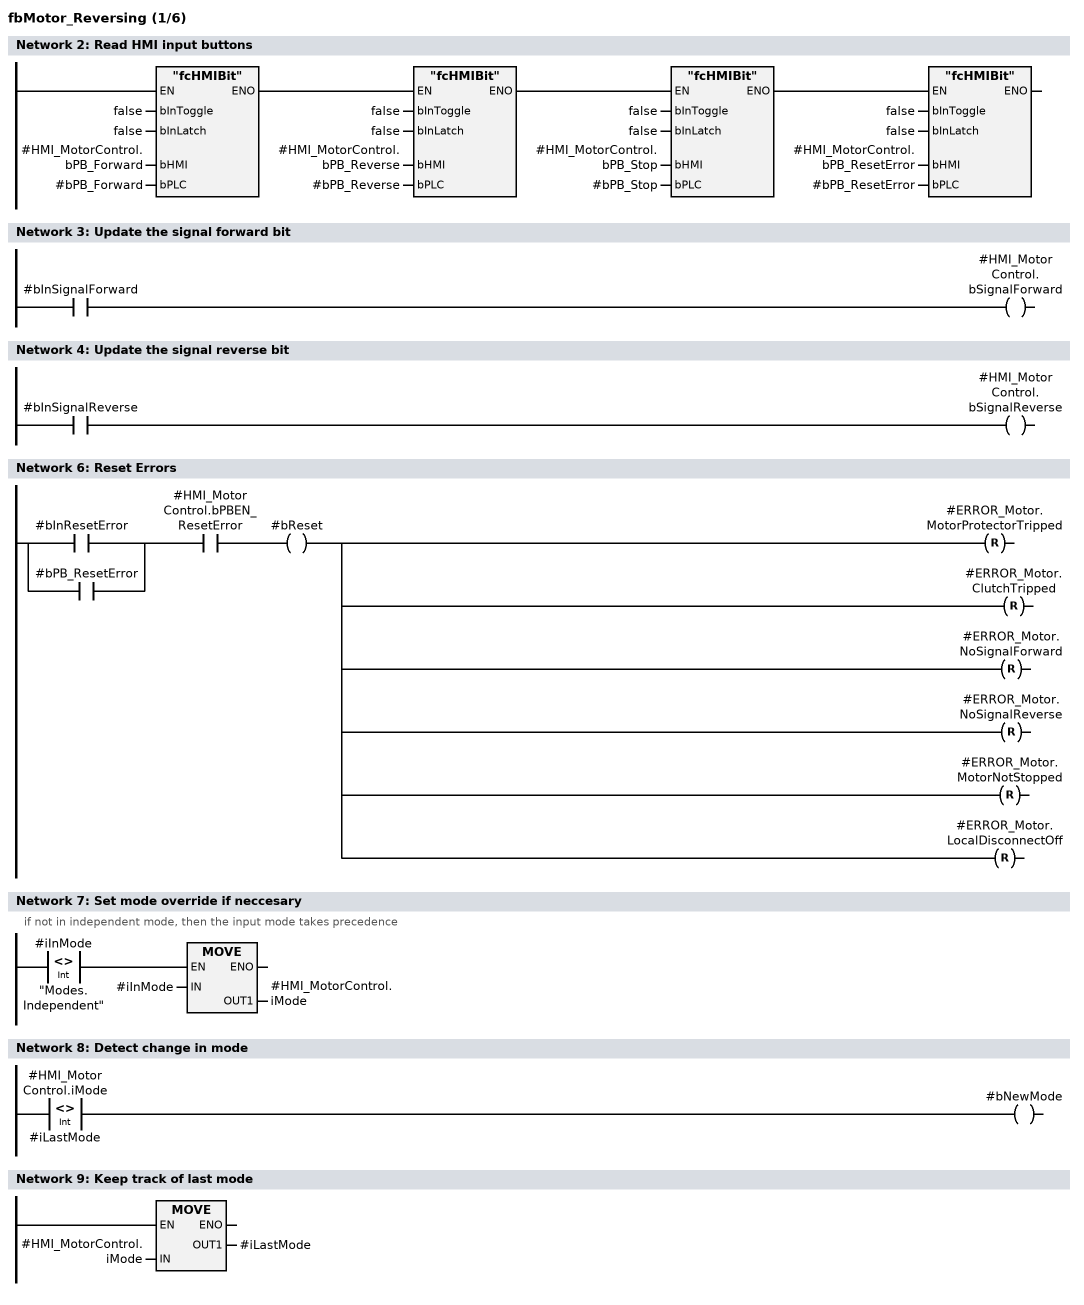
   RUNG wire#powerrail
      "fcHMIBit"(bInToggle := false, bInLatch := false, bHMI := #HMI_MotorControl.bPB_Forward, bPLC := #bPB_Forward)
      "fcHMIBit"(bInToggle := false, bInLatch := false, bHMI := #HMI_MotorControl.bPB_Reverse, bPLC := #bPB_Reverse)
      "fcHMIBit"(bInToggle := false, bInLatch := false, bHMI := #HMI_MotorControl.bPB_Stop, bPLC := #bPB_Stop)
      "fcHMIBit"(bInToggle := false, bInLatch := false, bHMI := #HMI_MotorControl.bPB_ResetError, bPLC := #bPB_ResetError)
   END_RUNG
   // the same network as SCL:
   "fcHMIBit"(bInToggle := false,
              bInLatch := false,
              bHMI := #HMI_MotorControl.bPB_Forward,
              bPLC := #bPB_Forward,
              ENO => #_w1);
   "fcHMIBit"(EN := #_w1,
              bInToggle := false,
              bInLatch := false,
              bHMI := #HMI_MotorControl.bPB_Reverse,
              bPLC := #bPB_Reverse,
              ENO => #_w2);
   "fcHMIBit"(EN := #_w2,
              bInToggle := false,
              bInLatch := false,
              bHMI := #HMI_MotorControl.bPB_Stop,
              bPLC := #bPB_Stop,
              ENO => #_w3);
   IF #_w3 THEN
       "fcHMIBit"(bInToggle := false,
                  bInLatch := false,
                  bHMI := #HMI_MotorControl.bPB_ResetError,
                  bPLC := #bPB_ResetError);
   END_IF;
END_REGION

REGION Network 3: Update the signal forward bit
   RUNG wire#powerrail
      Contact( #bInSignalForward )
      Coil( #HMI_MotorControl.bSignalForward )
   END_RUNG
   // the same network as SCL:
   #HMI_MotorControl.bSignalForward := #bInSignalForward;
END_REGION

REGION Network 4: Update the signal reverse bit
   RUNG wire#powerrail
      Contact( #bInSignalReverse )
      Coil( #HMI_MotorControl.bSignalReverse )
   END_RUNG
   // the same network as SCL:
   #HMI_MotorControl.bSignalReverse := #bInSignalReverse;
END_REGION

REGION Network 5: --------------------------------------------------- Control Logic ------------------------------------------------------------
END_REGION

REGION Network 6: Reset Errors
   RUNG wire#powerrail
      Contact( #bInResetError )
      wire#w1
      Contact( #HMI_MotorControl.bPBEN_ResetError )
      Coil( #bReset )
      wire#w2
      R_Coil( #ERROR_Motor.MotorProtectorTripped )
   END_RUNG
   RUNG wire#powerrail
      Contact( #bPB_ResetError )
   END_RUNG wire#w1
   RUNG wire#w2
      R_Coil( #ERROR_Motor.ClutchTripped )
   END_RUNG
   RUNG wire#w2
      R_Coil( #ERROR_Motor.NoSignalForward )
   END_RUNG
   RUNG wire#w2
      R_Coil( #ERROR_Motor.NoSignalReverse )
   END_RUNG
   RUNG wire#w2
      R_Coil( #ERROR_Motor.MotorNotStopped )
   END_RUNG
   RUNG wire#w2
      R_Coil( #ERROR_Motor.LocalDisconnectOff )
   END_RUNG
   // the same network as SCL:
   #bReset := (#bInResetError OR #bPB_ResetError) AND #HMI_MotorControl.bPBEN_ResetError;
   IF #bReset THEN
       #ERROR_Motor.MotorProtectorTripped := FALSE;
       #ERROR_Motor.ClutchTripped := FALSE;
       #ERROR_Motor.NoSignalForward := FALSE;
       #ERROR_Motor.NoSignalReverse := FALSE;
       #ERROR_Motor.MotorNotStopped := FALSE;
       #ERROR_Motor.LocalDisconnectOff := FALSE;
   END_IF;
END_REGION

REGION Network 7: Set mode override if neccesary
   // if not in independent mode, then the input mode takes precedence
   RUNG wire#powerrail
      { S7_Templates := "SrcType := Int" } NE_Contact(in1 := #iInMode, in2 := "Modes.Independent")
      { S7_GenerateENO := "TRUE" } Move(in := #iInMode, out1 => #HMI_MotorControl.iMode)
   END_RUNG
   // the same network as SCL:
   IF #iInMode <> "Modes.Independent" THEN #HMI_MotorControl.iMode := #iInMode; END_IF;
END_REGION

REGION Network 8: Detect change in mode
   RUNG wire#powerrail
      { S7_Templates := "SrcType := Int" } NE_Contact(in1 := #HMI_MotorControl.iMode, in2 := #iLastMode)
      Coil( #bNewMode )
   END_RUNG
   // the same network as SCL:
   #bNewMode := #HMI_MotorControl.iMode <> #iLastMode;
END_REGION

REGION Network 9: Keep track of last mode
   RUNG wire#powerrail
      { S7_GenerateENO := "TRUE" } Move(in := #HMI_MotorControl.iMode, out1 => #iLastMode)
   END_RUNG
   // the same network as SCL:
   #iLastMode := #HMI_MotorControl.iMode;
END_REGION

REGION Network 10: Determine if auto or manual mode is active
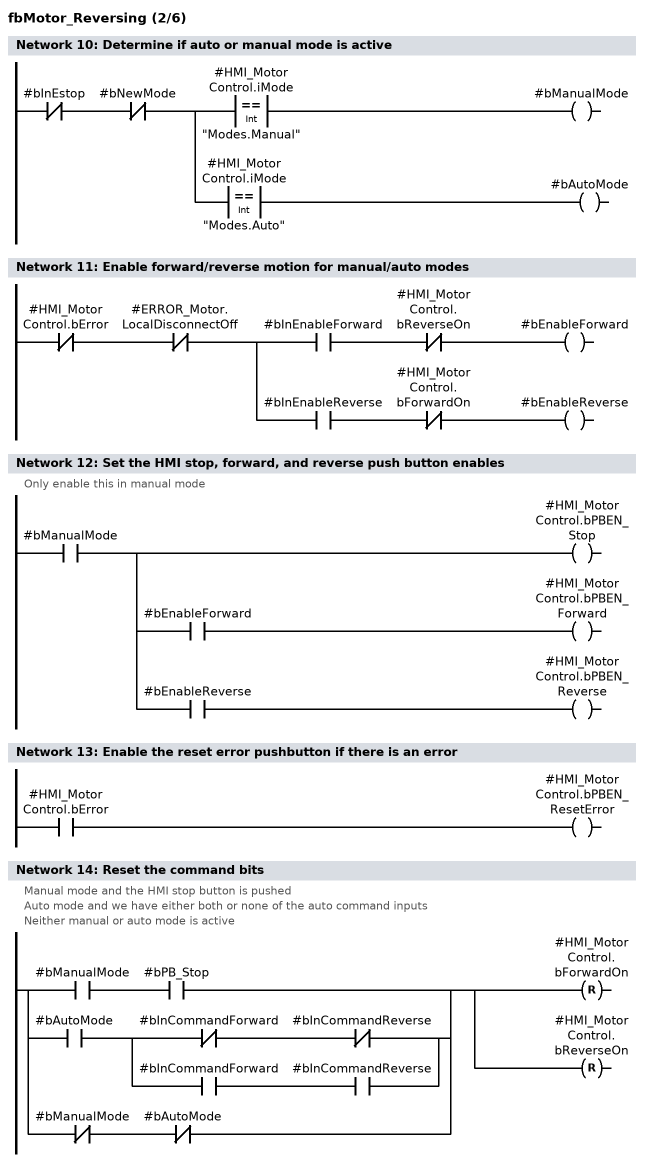
   RUNG wire#powerrail
      I_Contact( #bInEstop )
      I_Contact( #bNewMode )
      wire#w1
      { S7_Templates := "SrcType := Int" } EQ_Contact(in1 := #HMI_MotorControl.iMode, in2 := "Modes.Manual")
      Coil( #bManualMode )
   END_RUNG
   RUNG wire#w1
      { S7_Templates := "SrcType := Int" } EQ_Contact(in1 := #HMI_MotorControl.iMode, in2 := "Modes.Auto")
      Coil( #bAutoMode )
   END_RUNG
   // the same network as SCL:
   #_w1 := NOT #bInEstop AND NOT #bNewMode;
   #bManualMode := #_w1 AND (#HMI_MotorControl.iMode = "Modes.Manual");
   #bAutoMode := #_w1 AND (#HMI_MotorControl.iMode = "Modes.Auto");
END_REGION

REGION Network 11: Enable forward/reverse motion for manual/auto modes
   RUNG wire#powerrail
      I_Contact( #HMI_MotorControl.bError )
      I_Contact( #ERROR_Motor.LocalDisconnectOff )
      wire#w1
      Contact( #bInEnableForward )
      I_Contact( #HMI_MotorControl.bReverseOn )
      Coil( #bEnableForward )
   END_RUNG
   RUNG wire#w1
      Contact( #bInEnableReverse )
      I_Contact( #HMI_MotorControl.bForwardOn )
      Coil( #bEnableReverse )
   END_RUNG
   // the same network as SCL:
   #_w1 := NOT #HMI_MotorControl.bError AND NOT #ERROR_Motor.LocalDisconnectOff;
   #bEnableForward := #_w1 AND #bInEnableForward AND NOT #HMI_MotorControl.bReverseOn;
   #bEnableReverse := #_w1 AND #bInEnableReverse AND NOT #HMI_MotorControl.bForwardOn;
END_REGION

REGION Network 12: Set the HMI stop, forward, and reverse push button enables
   // Only enable this in manual mode
   RUNG wire#powerrail
      Contact( #bManualMode )
      wire#w1
      Coil( #HMI_MotorControl.bPBEN_Stop )
   END_RUNG
   RUNG wire#w1
      Contact( #bEnableForward )
      Coil( #HMI_MotorControl.bPBEN_Forward )
   END_RUNG
   RUNG wire#w1
      Contact( #bEnableReverse )
      Coil( #HMI_MotorControl.bPBEN_Reverse )
   END_RUNG
   // the same network as SCL:
   #HMI_MotorControl.bPBEN_Stop := #bManualMode;
   #HMI_MotorControl.bPBEN_Forward := #bManualMode AND #bEnableForward;
   #HMI_MotorControl.bPBEN_Reverse := #bManualMode AND #bEnableReverse;
END_REGION

REGION Network 13: Enable the reset error pushbutton if there is an error
   RUNG wire#powerrail
      Contact( #HMI_MotorControl.bError )
      Coil( #HMI_MotorControl.bPBEN_ResetError )
   END_RUNG
   // the same network as SCL:
   #HMI_MotorControl.bPBEN_ResetError := #HMI_MotorControl.bError;
END_REGION

REGION Network 14: Reset the command bits
   // Manual mode and the HMI stop button is pushed
   // Auto mode and we have either both or none of the auto command inputs
   // Neither manual or auto mode is active
   RUNG wire#powerrail
      Contact( #bManualMode )
      Contact( #bPB_Stop )
      wire#w1
      R_Coil( #HMI_MotorControl.bForwardOn )
   END_RUNG
   RUNG wire#powerrail
      Contact( #bAutoMode )
      wire#w2
      I_Contact( #bInCommandForward )
      I_Contact( #bInCommandReverse )
   END_RUNG wire#w1
   RUNG wire#w2
      Contact( #bInCommandForward )
      Contact( #bInCommandReverse )
   END_RUNG wire#w1
   RUNG wire#powerrail
      I_Contact( #bManualMode )
      I_Contact( #bAutoMode )
   END_RUNG wire#w1
   RUNG wire#w1
      R_Coil( #HMI_MotorControl.bReverseOn )
   END_RUNG
   // the same network as SCL:
   IF (#bManualMode AND #bPB_Stop) OR (#bAutoMode AND ((NOT #bInCommandForward AND NOT #bInCommandReverse) OR (#bInCommandForward AND #bInCommandReverse))) OR (NOT #bManualMode AND NOT #bAutoMode) THEN
       #HMI_MotorControl.bForwardOn := FALSE;
       #HMI_MotorControl.bReverseOn := FALSE;
   END_IF;
END_REGION

REGION Network 15: Start forward request
   // Manual mode and only a start forward button is pressed and enabled
   // Auto mode when we receive a auto command and it is enabled
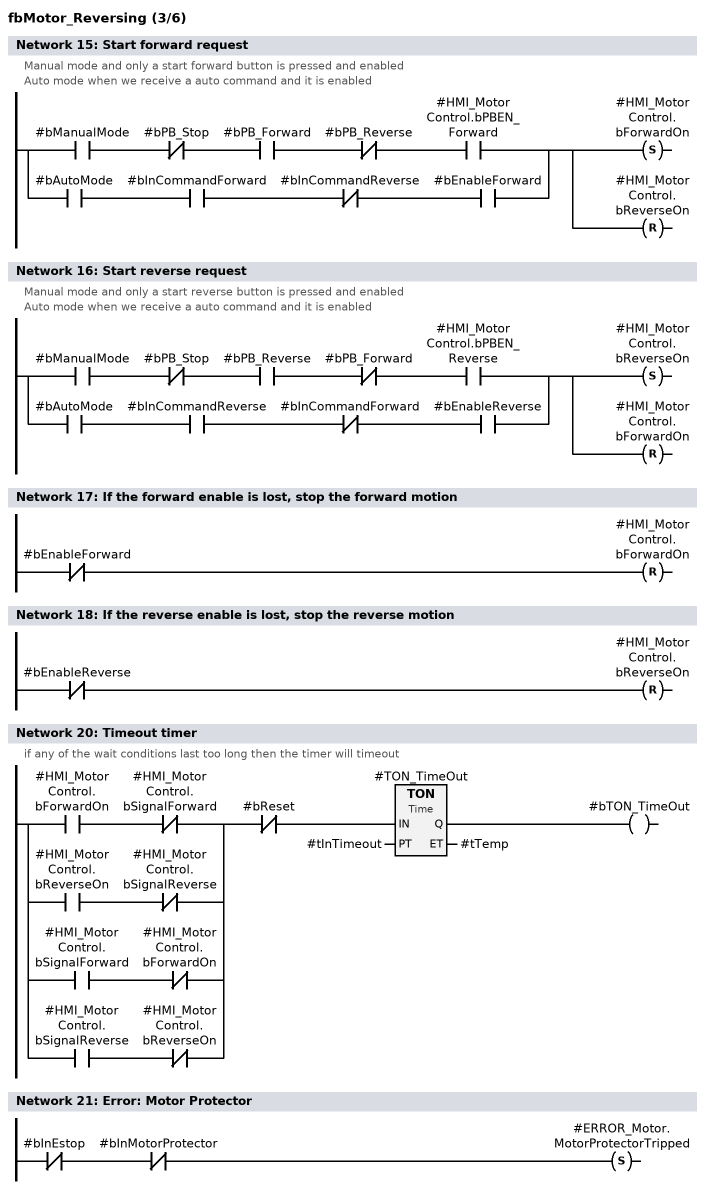
   RUNG wire#powerrail
      Contact( #bManualMode )
      I_Contact( #bPB_Stop )
      Contact( #bPB_Forward )
      I_Contact( #bPB_Reverse )
      Contact( #HMI_MotorControl.bPBEN_Forward )
      wire#w1
      S_Coil( #HMI_MotorControl.bForwardOn )
   END_RUNG
   RUNG wire#powerrail
      Contact( #bAutoMode )
      Contact( #bInCommandForward )
      I_Contact( #bInCommandReverse )
      Contact( #bEnableForward )
   END_RUNG wire#w1
   RUNG wire#w1
      R_Coil( #HMI_MotorControl.bReverseOn )
   END_RUNG
   // the same network as SCL:
   IF (#bManualMode AND NOT #bPB_Stop AND #bPB_Forward AND NOT #bPB_Reverse AND #HMI_MotorControl.bPBEN_Forward) OR (#bAutoMode AND #bInCommandForward AND NOT #bInCommandReverse AND #bEnableForward) THEN
       #HMI_MotorControl.bForwardOn := TRUE;
       #HMI_MotorControl.bReverseOn := FALSE;
   END_IF;
END_REGION

REGION Network 16: Start reverse request
   // Manual mode and only a start reverse button is pressed and enabled
   // Auto mode when we receive a auto command and it is enabled
   RUNG wire#powerrail
      Contact( #bManualMode )
      I_Contact( #bPB_Stop )
      Contact( #bPB_Reverse )
      I_Contact( #bPB_Forward )
      Contact( #HMI_MotorControl.bPBEN_Reverse )
      wire#w1
      S_Coil( #HMI_MotorControl.bReverseOn )
   END_RUNG
   RUNG wire#powerrail
      Contact( #bAutoMode )
      Contact( #bInCommandReverse )
      I_Contact( #bInCommandForward )
      Contact( #bEnableReverse )
   END_RUNG wire#w1
   RUNG wire#w1
      R_Coil( #HMI_MotorControl.bForwardOn )
   END_RUNG
   // the same network as SCL:
   IF (#bManualMode AND NOT #bPB_Stop AND #bPB_Reverse AND NOT #bPB_Forward AND #HMI_MotorControl.bPBEN_Reverse) OR (#bAutoMode AND #bInCommandReverse AND NOT #bInCommandForward AND #bEnableReverse) THEN
       #HMI_MotorControl.bReverseOn := TRUE;
       #HMI_MotorControl.bForwardOn := FALSE;
   END_IF;
END_REGION

REGION Network 17: If the forward enable is lost, stop the forward motion
   RUNG wire#powerrail
      I_Contact( #bEnableForward )
      R_Coil( #HMI_MotorControl.bForwardOn )
   END_RUNG
   // the same network as SCL:
   IF NOT #bEnableForward THEN #HMI_MotorControl.bForwardOn := FALSE; END_IF;
END_REGION

REGION Network 18: If the reverse enable is lost, stop the reverse motion
   RUNG wire#powerrail
      I_Contact( #bEnableReverse )
      R_Coil( #HMI_MotorControl.bReverseOn )
   END_RUNG
   // the same network as SCL:
   IF NOT #bEnableReverse THEN #HMI_MotorControl.bReverseOn := FALSE; END_IF;
END_REGION

REGION Network 19: --------------------------------------------------------- Errors ------------------------------------------------------------------
END_REGION

REGION Network 20: Timeout timer
   // if any of the wait conditions last too long then the timer will timeout
   #TON_TimeOut.TON(IN := ((#HMI_MotorControl.bForwardOn AND NOT #HMI_MotorControl.bSignalForward) OR (#HMI_MotorControl.bReverseOn AND NOT #HMI_MotorControl.bSignalReverse) OR (#HMI_MotorControl.bSignalForward AND NOT #HMI_MotorControl.bForwardOn) OR (#HMI_MotorControl.bSignalReverse AND NOT #HMI_MotorControl.bReverseOn)) AND NOT #bReset,
                    PT := #tInTimeout,
                    ET => #tTemp);
   #bTON_TimeOut := #TON_TimeOut.Q;
END_REGION

REGION Network 21: Error: Motor Protector
   RUNG wire#powerrail
      I_Contact( #bInEstop )
      I_Contact( #bInMotorProtector )
      S_Coil( #ERROR_Motor.MotorProtectorTripped )
   END_RUNG
   // the same network as SCL:
   IF NOT #bInEstop AND NOT #bInMotorProtector THEN #ERROR_Motor.MotorProtectorTripped := TRUE; END_IF;
END_REGION

REGION Network 22: Error: Kill Switch/ local disconnect
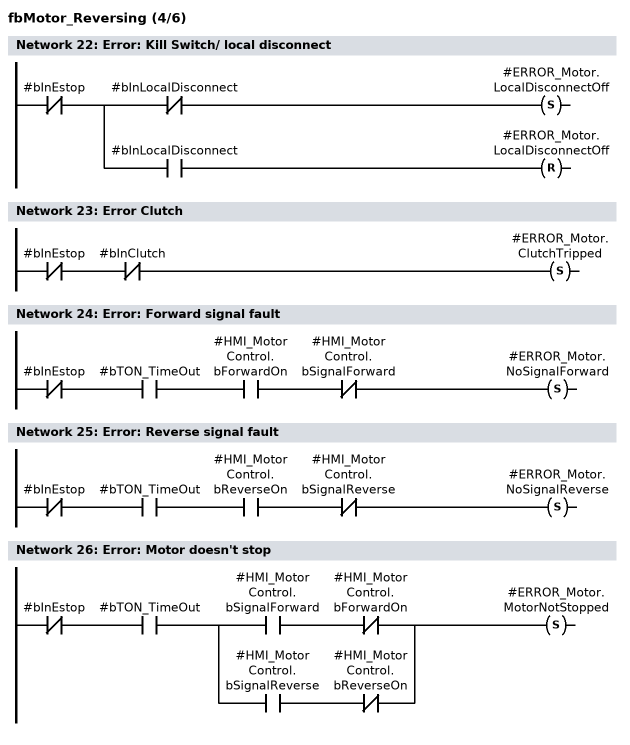
   RUNG wire#powerrail
      I_Contact( #bInEstop )
      wire#w1
      I_Contact( #bInLocalDisconnect )
      S_Coil( #ERROR_Motor.LocalDisconnectOff )
   END_RUNG
   RUNG wire#w1
      Contact( #bInLocalDisconnect )
      R_Coil( #ERROR_Motor.LocalDisconnectOff )
   END_RUNG
   // the same network as SCL:
   IF NOT #bInEstop AND NOT #bInLocalDisconnect THEN #ERROR_Motor.LocalDisconnectOff := TRUE; END_IF;
   IF NOT #bInEstop AND #bInLocalDisconnect THEN #ERROR_Motor.LocalDisconnectOff := FALSE; END_IF;
END_REGION

REGION Network 23: Error Clutch
   RUNG wire#powerrail
      I_Contact( #bInEstop )
      I_Contact( #bInClutch )
      S_Coil( #ERROR_Motor.ClutchTripped )
   END_RUNG
   // the same network as SCL:
   IF NOT #bInEstop AND NOT #bInClutch THEN #ERROR_Motor.ClutchTripped := TRUE; END_IF;
END_REGION

REGION Network 24: Error: Forward signal fault
   RUNG wire#powerrail
      I_Contact( #bInEstop )
      Contact( #bTON_TimeOut )
      Contact( #HMI_MotorControl.bForwardOn )
      I_Contact( #HMI_MotorControl.bSignalForward )
      S_Coil( #ERROR_Motor.NoSignalForward )
   END_RUNG
   // the same network as SCL:
   IF NOT #bInEstop AND #bTON_TimeOut AND #HMI_MotorControl.bForwardOn AND NOT #HMI_MotorControl.bSignalForward THEN
       #ERROR_Motor.NoSignalForward := TRUE;
   END_IF;
END_REGION

REGION Network 25: Error: Reverse signal fault
   RUNG wire#powerrail
      I_Contact( #bInEstop )
      Contact( #bTON_TimeOut )
      Contact( #HMI_MotorControl.bReverseOn )
      I_Contact( #HMI_MotorControl.bSignalReverse )
      S_Coil( #ERROR_Motor.NoSignalReverse )
   END_RUNG
   // the same network as SCL:
   IF NOT #bInEstop AND #bTON_TimeOut AND #HMI_MotorControl.bReverseOn AND NOT #HMI_MotorControl.bSignalReverse THEN
       #ERROR_Motor.NoSignalReverse := TRUE;
   END_IF;
END_REGION

REGION Network 26: Error: Motor doesn't stop
   RUNG wire#powerrail
      I_Contact( #bInEstop )
      Contact( #bTON_TimeOut )
      wire#w1
      Contact( #HMI_MotorControl.bSignalForward )
      I_Contact( #HMI_MotorControl.bForwardOn )
      wire#w2
      S_Coil( #ERROR_Motor.MotorNotStopped )
   END_RUNG
   RUNG wire#w1
      Contact( #HMI_MotorControl.bSignalReverse )
      I_Contact( #HMI_MotorControl.bReverseOn )
   END_RUNG wire#w2
   // the same network as SCL:
   IF NOT #bInEstop AND #bTON_TimeOut AND ((#HMI_MotorControl.bSignalForward AND NOT #HMI_MotorControl.bForwardOn) OR (#HMI_MotorControl.bSignalReverse AND NOT #HMI_MotorControl.bReverseOn)) THEN
       #ERROR_Motor.MotorNotStopped := TRUE;
   END_IF;
END_REGION

REGION Network 27: Scroll errors on the HMI
   // This block loops through all of the possible erros and displays them on the HMI 
   // by setting an index value for each error bit.
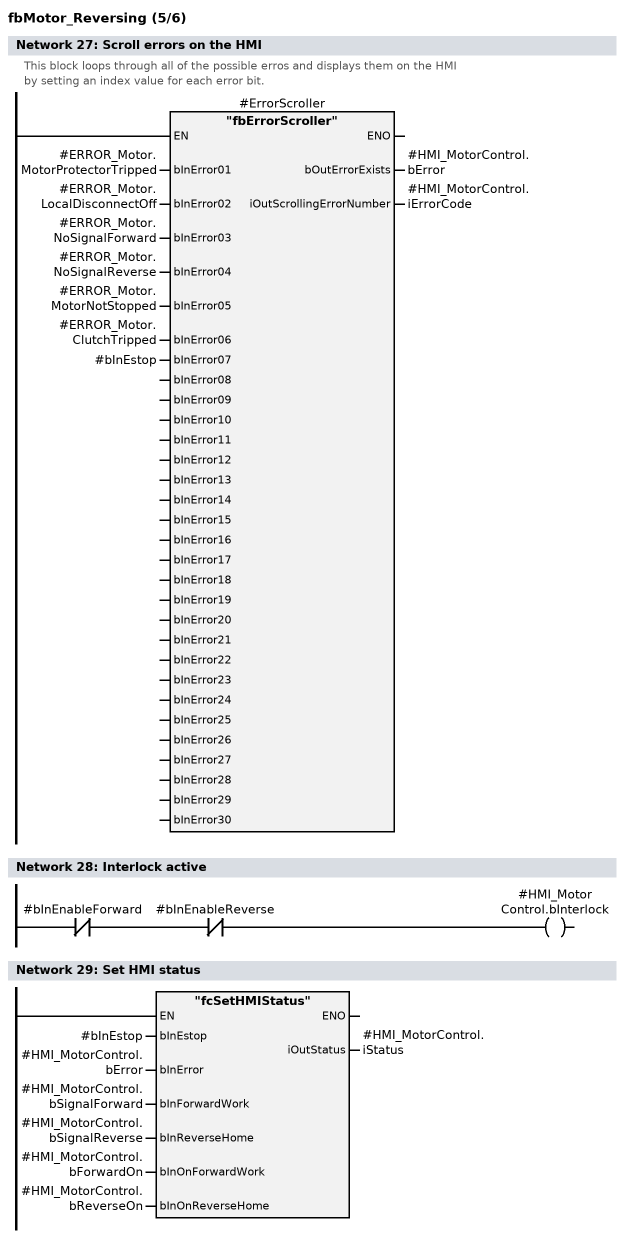
   RUNG wire#powerrail
      #ErrorScroller(bInError01 := #ERROR_Motor.MotorProtectorTripped, bInError02 := #ERROR_Motor.LocalDisconnectOff, bInError03 := #ERROR_Motor.NoSignalForward, bInError04 := #ERROR_Motor.NoSignalReverse, bInError05 := #ERROR_Motor.MotorNotStopped, bInError06 := #ERROR_Motor.ClutchTripped, bInError07 := #bInEstop, bInError08 :=, bInError09 :=, bInError10 :=, bInError11 :=, bInError12 :=, bInError13 :=, bInError14 :=, bInError15 :=, bInError16 :=, bInError17 :=, bInError18 :=, bInError19 :=, bInError20 :=, bInError21 :=, bInError22 :=, bInError23 :=, bInError24 :=, bInError25 :=, bInError26 :=, bInError27 :=, bInError28 :=, bInError29 :=, bInError30 :=, bOutErrorExists => #HMI_MotorControl.bError, iOutScrollingErrorNumber => #HMI_MotorControl.iErrorCode)
   END_RUNG
   // the same network as SCL:
   #ErrorScroller(bInError01 := #ERROR_Motor.MotorProtectorTripped,   // "fbErrorScroller"
                  bInError02 := #ERROR_Motor.LocalDisconnectOff,
                  bInError03 := #ERROR_Motor.NoSignalForward,
                  bInError04 := #ERROR_Motor.NoSignalReverse,
                  bInError05 := #ERROR_Motor.MotorNotStopped,
                  bInError06 := #ERROR_Motor.ClutchTripped,
                  bInError07 := #bInEstop,
                  bOutErrorExists => #HMI_MotorControl.bError,
                  iOutScrollingErrorNumber => #HMI_MotorControl.iErrorCode);
END_REGION

REGION Network 28: Interlock active
   RUNG wire#powerrail
      I_Contact( #bInEnableForward )
      I_Contact( #bInEnableReverse )
      Coil( #HMI_MotorControl.bInterlock )
   END_RUNG
   // the same network as SCL:
   #HMI_MotorControl.bInterlock := NOT #bInEnableForward AND NOT #bInEnableReverse;
END_REGION

REGION Network 29: Set HMI status
   RUNG wire#powerrail
      "fcSetHMIStatus"(bInEstop := #bInEstop, bInError := #HMI_MotorControl.bError, bInForwardWork := #HMI_MotorControl.bSignalForward, bInReverseHome := #HMI_MotorControl.bSignalReverse, bInOnForwardWork := #HMI_MotorControl.bForwardOn, bInOnReverseHome := #HMI_MotorControl.bReverseOn, iOutStatus => #HMI_MotorControl.iStatus)
   END_RUNG
   // the same network as SCL:
   "fcSetHMIStatus"(bInEstop := #bInEstop,
                    bInError := #HMI_MotorControl.bError,
                    bInForwardWork := #HMI_MotorControl.bSignalForward,
                    bInReverseHome := #HMI_MotorControl.bSignalReverse,
                    bInOnForwardWork := #HMI_MotorControl.bForwardOn,
                    bInOnReverseHome := #HMI_MotorControl.bReverseOn,
                    iOutStatus => #HMI_MotorControl.iStatus);
END_REGION

REGION Network 30: ------------------------------------------------- Outputs --------------------------------------------------
END_REGION

REGION Network 31: Output: Forward
   // Forward
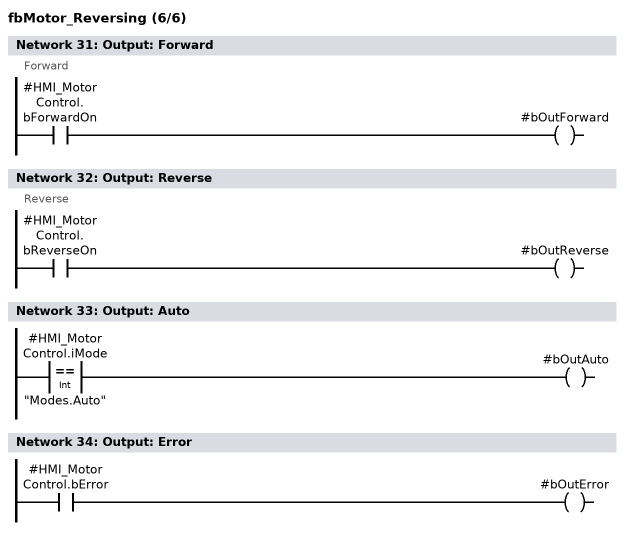
   RUNG wire#powerrail
      Contact( #HMI_MotorControl.bForwardOn )
      Coil( #bOutForward )
   END_RUNG
   // the same network as SCL:
   #bOutForward := #HMI_MotorControl.bForwardOn;
END_REGION

REGION Network 32: Output: Reverse
   // Reverse
   RUNG wire#powerrail
      Contact( #HMI_MotorControl.bReverseOn )
      Coil( #bOutReverse )
   END_RUNG
   // the same network as SCL:
   #bOutReverse := #HMI_MotorControl.bReverseOn;
END_REGION

REGION Network 33: Output: Auto
   RUNG wire#powerrail
      { S7_Templates := "SrcType := Int" } EQ_Contact(in1 := #HMI_MotorControl.iMode, in2 := "Modes.Auto")
      Coil( #bOutAuto )
   END_RUNG
   // the same network as SCL:
   #bOutAuto := #HMI_MotorControl.iMode = "Modes.Auto";
END_REGION

REGION Network 34: Output: Error
   RUNG wire#powerrail
      Contact( #HMI_MotorControl.bError )
      Coil( #bOutError )
   END_RUNG
   // the same network as SCL:
   #bOutError := #HMI_MotorControl.bError;
END_REGION
END_FUNCTION_BLOCK

FUNCTION_BLOCK "fbIO_AnalogInput"   // FB140, LAD
TITLE = Reads and controls an analog input
{ S7_Optimized_Access := 'FALSE' }
VERSION : 0.1
BEGIN

REGION Network 1: --------------------------------------------------------- Inputs ------------------------------------------------------------------
END_REGION

REGION Network 2: Read HMI input buttons
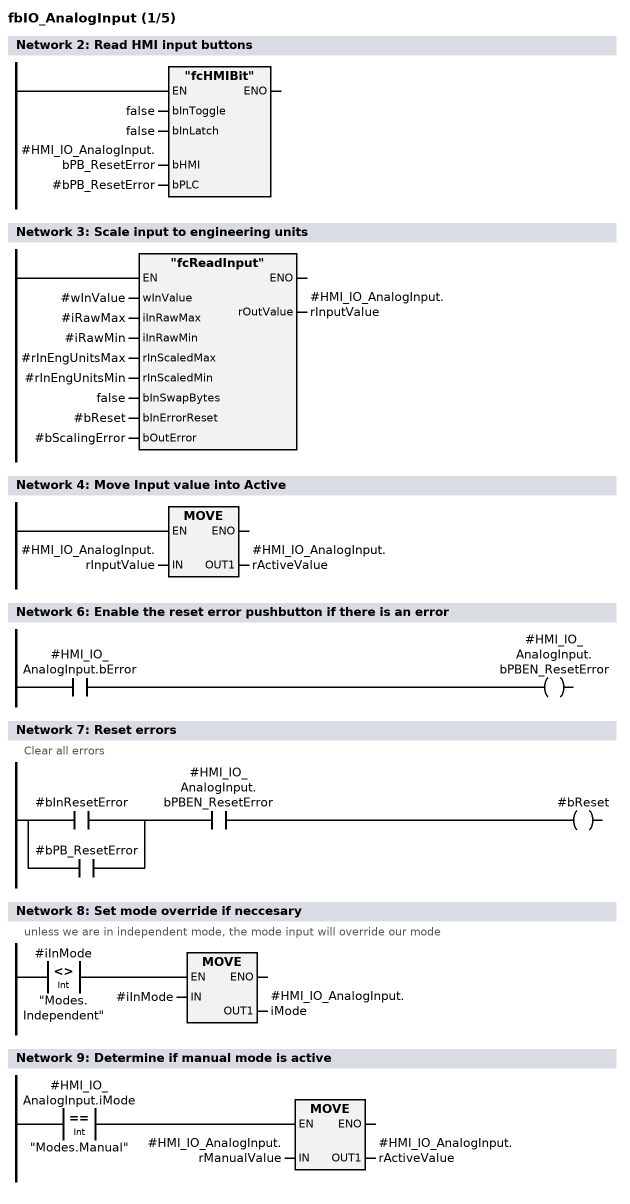
   RUNG wire#powerrail
      "fcHMIBit"(bInToggle := false, bInLatch := false, bHMI := #HMI_IO_AnalogInput.bPB_ResetError, bPLC := #bPB_ResetError)
   END_RUNG
   // the same network as SCL:
   "fcHMIBit"(bInToggle := false,
              bInLatch := false,
              bHMI := #HMI_IO_AnalogInput.bPB_ResetError,
              bPLC := #bPB_ResetError);
END_REGION

REGION Network 3: Scale input to engineering units
   RUNG wire#powerrail
      "fcReadInput"(wInValue := #wInValue, iInRawMax := #iRawMax, iInRawMin := #iRawMin, rInScaledMax := #rInEngUnitsMax, rInScaledMin := #rInEngUnitsMin, bInSwapBytes := false, bInErrorReset := #bReset, bOutError := #bScalingError, rOutValue => #HMI_IO_AnalogInput.rInputValue)
   END_RUNG
   // the same network as SCL:
   "fcReadInput"(wInValue := #wInValue,
                 iInRawMax := #iRawMax,
                 iInRawMin := #iRawMin,
                 rInScaledMax := #rInEngUnitsMax,
                 rInScaledMin := #rInEngUnitsMin,
                 bInSwapBytes := false,
                 bInErrorReset := #bReset,
                 bOutError := #bScalingError,
                 rOutValue => #HMI_IO_AnalogInput.rInputValue);
END_REGION

REGION Network 4: Move Input value into Active
   RUNG wire#powerrail
      Move(in := #HMI_IO_AnalogInput.rInputValue, out1 => #HMI_IO_AnalogInput.rActiveValue)
   END_RUNG
   // the same network as SCL:
   #HMI_IO_AnalogInput.rActiveValue := #HMI_IO_AnalogInput.rInputValue;
END_REGION

REGION Network 5: --------------------------------------------------- Control Logic ------------------------------------------------------------
END_REGION

REGION Network 6: Enable the reset error pushbutton if there is an error
   RUNG wire#powerrail
      Contact( #HMI_IO_AnalogInput.bError )
      Coil( #HMI_IO_AnalogInput.bPBEN_ResetError )
   END_RUNG
   // the same network as SCL:
   #HMI_IO_AnalogInput.bPBEN_ResetError := #HMI_IO_AnalogInput.bError;
END_REGION

REGION Network 7: Reset errors
   // Clear all errors
   RUNG wire#powerrail
      Contact( #bInResetError )
      wire#w1
      Contact( #HMI_IO_AnalogInput.bPBEN_ResetError )
      Coil( #bReset )
   END_RUNG
   RUNG wire#powerrail
      Contact( #bPB_ResetError )
   END_RUNG wire#w1
   // the same network as SCL:
   #bReset := (#bInResetError OR #bPB_ResetError) AND #HMI_IO_AnalogInput.bPBEN_ResetError;
END_REGION

REGION Network 8: Set mode override if neccesary
   // unless we are in independent mode, the mode input will override our mode
   RUNG wire#powerrail
      { S7_Templates := "SrcType := Int" } NE_Contact(in1 := #iInMode, in2 := "Modes.Independent")
      { S7_GenerateENO := "TRUE" } Move(in := #iInMode, out1 => #HMI_IO_AnalogInput.iMode)
   END_RUNG
   // the same network as SCL:
   IF #iInMode <> "Modes.Independent" THEN #HMI_IO_AnalogInput.iMode := #iInMode; END_IF;
END_REGION

REGION Network 9: Determine if manual mode is active
   RUNG wire#powerrail
      { S7_Templates := "SrcType := Int" } EQ_Contact(in1 := #HMI_IO_AnalogInput.iMode, in2 := "Modes.Manual")
      { S7_GenerateENO := "TRUE" } Move(in := #HMI_IO_AnalogInput.rManualValue, out1 => #HMI_IO_AnalogInput.rActiveValue)
   END_RUNG
   // the same network as SCL:
   IF #HMI_IO_AnalogInput.iMode = "Modes.Manual" THEN
       #HMI_IO_AnalogInput.rActiveValue := #HMI_IO_AnalogInput.rManualValue;
   END_IF;
END_REGION

REGION Network 10: Default sensor type
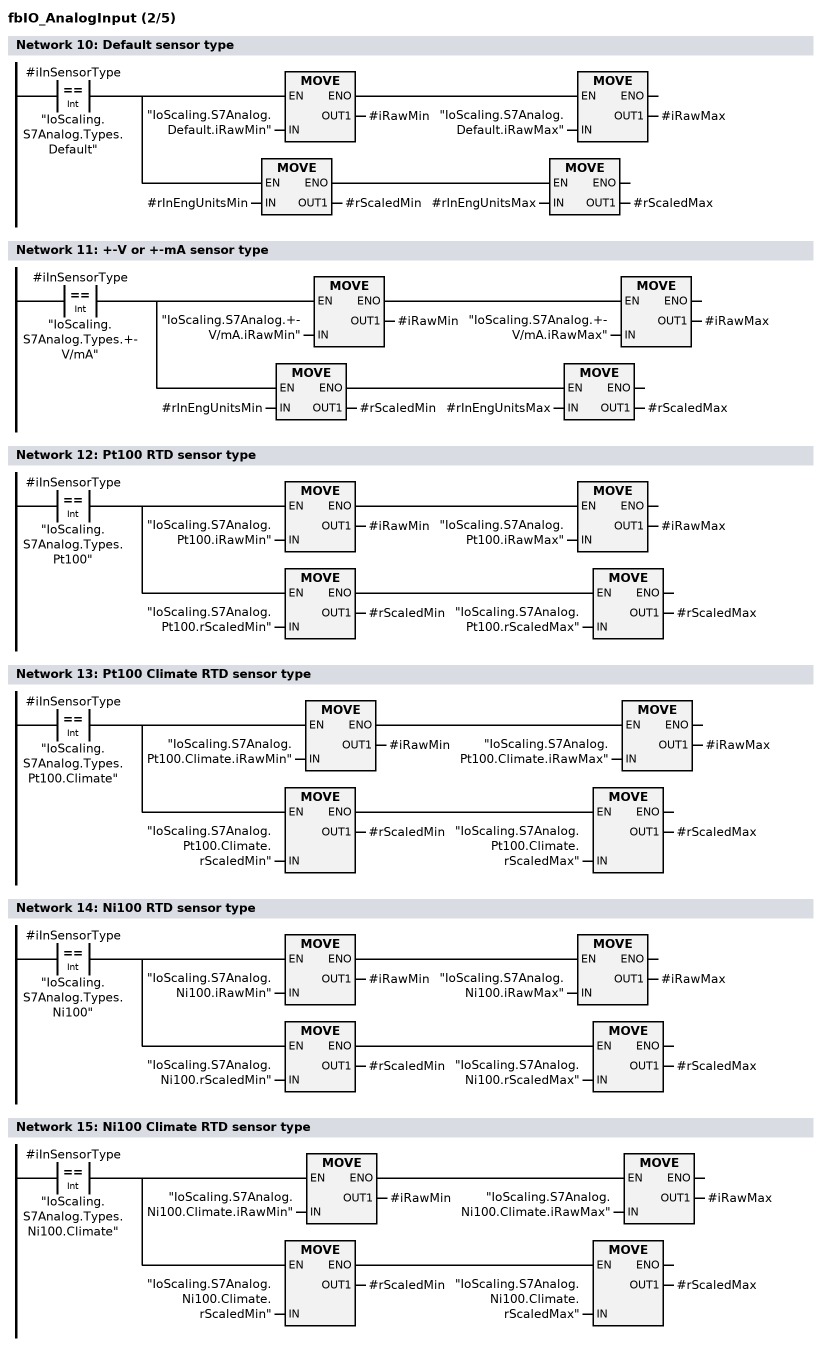
   RUNG wire#powerrail
      { S7_Templates := "SrcType := Int" } EQ_Contact(in1 := #iInSensorType, in2 := "IoScaling.S7Analog.Types.Default")
      wire#w1
      { S7_GenerateENO := "TRUE" } Move(in := "IoScaling.S7Analog.Default.iRawMin", out1 => #iRawMin)
      { S7_GenerateENO := "TRUE" } Move(in := "IoScaling.S7Analog.Default.iRawMax", out1 => #iRawMax)
   END_RUNG
   RUNG wire#w1
      { S7_GenerateENO := "TRUE" } Move(in := #rInEngUnitsMin, out1 => #rScaledMin)
      { S7_GenerateENO := "TRUE" } Move(in := #rInEngUnitsMax, out1 => #rScaledMax)
   END_RUNG
   // the same network as SCL:
   // ENO of a box is taken as its EN; it also drops when the box reports an error
   IF #iInSensorType = "IoScaling.S7Analog.Types.Default" THEN
       #iRawMin := "IoScaling.S7Analog.Default.iRawMin";
       #iRawMax := "IoScaling.S7Analog.Default.iRawMax";
       #rScaledMin := #rInEngUnitsMin;
       #rScaledMax := #rInEngUnitsMax;
   END_IF;
END_REGION

REGION Network 11: +-V or +-mA sensor type
   RUNG wire#powerrail
      { S7_Templates := "SrcType := Int" } EQ_Contact(in1 := #iInSensorType, in2 := "IoScaling.S7Analog.Types.+-V/mA")
      wire#w1
      { S7_GenerateENO := "TRUE" } Move(in := "IoScaling.S7Analog.+-V/mA.iRawMin", out1 => #iRawMin)
      { S7_GenerateENO := "TRUE" } Move(in := "IoScaling.S7Analog.+-V/mA.iRawMax", out1 => #iRawMax)
   END_RUNG
   RUNG wire#w1
      { S7_GenerateENO := "TRUE" } Move(in := #rInEngUnitsMin, out1 => #rScaledMin)
      { S7_GenerateENO := "TRUE" } Move(in := #rInEngUnitsMax, out1 => #rScaledMax)
   END_RUNG
   // the same network as SCL:
   // ENO of a box is taken as its EN; it also drops when the box reports an error
   IF #iInSensorType = "IoScaling.S7Analog.Types.+-V/mA" THEN
       #iRawMin := "IoScaling.S7Analog.+-V/mA.iRawMin";
       #iRawMax := "IoScaling.S7Analog.+-V/mA.iRawMax";
       #rScaledMin := #rInEngUnitsMin;
       #rScaledMax := #rInEngUnitsMax;
   END_IF;
END_REGION

REGION Network 12: Pt100 RTD sensor type
   RUNG wire#powerrail
      { S7_Templates := "SrcType := Int" } EQ_Contact(in1 := #iInSensorType, in2 := "IoScaling.S7Analog.Types.Pt100")
      wire#w1
      { S7_GenerateENO := "TRUE" } Move(in := "IoScaling.S7Analog.Pt100.iRawMin", out1 => #iRawMin)
      { S7_GenerateENO := "TRUE" } Move(in := "IoScaling.S7Analog.Pt100.iRawMax", out1 => #iRawMax)
   END_RUNG
   RUNG wire#w1
      { S7_GenerateENO := "TRUE" } Move(in := "IoScaling.S7Analog.Pt100.rScaledMin", out1 => #rScaledMin)
      { S7_GenerateENO := "TRUE" } Move(in := "IoScaling.S7Analog.Pt100.rScaledMax", out1 => #rScaledMax)
   END_RUNG
   // the same network as SCL:
   // ENO of a box is taken as its EN; it also drops when the box reports an error
   IF #iInSensorType = "IoScaling.S7Analog.Types.Pt100" THEN
       #iRawMin := "IoScaling.S7Analog.Pt100.iRawMin";
       #iRawMax := "IoScaling.S7Analog.Pt100.iRawMax";
       #rScaledMin := "IoScaling.S7Analog.Pt100.rScaledMin";
       #rScaledMax := "IoScaling.S7Analog.Pt100.rScaledMax";
   END_IF;
END_REGION

REGION Network 13: Pt100 Climate RTD sensor type
   RUNG wire#powerrail
      { S7_Templates := "SrcType := Int" } EQ_Contact(in1 := #iInSensorType, in2 := "IoScaling.S7Analog.Types.Pt100.Climate")
      wire#w1
      { S7_GenerateENO := "TRUE" } Move(in := "IoScaling.S7Analog.Pt100.Climate.iRawMin", out1 => #iRawMin)
      { S7_GenerateENO := "TRUE" } Move(in := "IoScaling.S7Analog.Pt100.Climate.iRawMax", out1 => #iRawMax)
   END_RUNG
   RUNG wire#w1
      { S7_GenerateENO := "TRUE" } Move(in := "IoScaling.S7Analog.Pt100.Climate.rScaledMin", out1 => #rScaledMin)
      { S7_GenerateENO := "TRUE" } Move(in := "IoScaling.S7Analog.Pt100.Climate.rScaledMax", out1 => #rScaledMax)
   END_RUNG
   // the same network as SCL:
   // ENO of a box is taken as its EN; it also drops when the box reports an error
   IF #iInSensorType = "IoScaling.S7Analog.Types.Pt100.Climate" THEN
       #iRawMin := "IoScaling.S7Analog.Pt100.Climate.iRawMin";
       #iRawMax := "IoScaling.S7Analog.Pt100.Climate.iRawMax";
       #rScaledMin := "IoScaling.S7Analog.Pt100.Climate.rScaledMin";
       #rScaledMax := "IoScaling.S7Analog.Pt100.Climate.rScaledMax";
   END_IF;
END_REGION